(* Logix 5000 project; controller MV vendor 1 type 14 code 217 rev 31.11; software revision 31.00; part 46 of 53 *)
(* tags used below, declared in another part *)
   Always_Off : BOOL;
   CWD : CHECKWORD_FLAGS;
   Enable_TimeString : BOOL;
   MC_N100 : INT[255];   // C1_PLC Channel 1 PLC data
   MC_N120 : INT[255];   // C2 PLC Channel 2 PLC data
   MV_BM01_AV01 : PlantItem;   // BM01_AV01
   MV_BM01_AV01_CIP : BOOL;
   MV_BM01_AV01_mv22 : BOOL;
   MV_BM01_ZS04 : PlantItem;   // BM01ZS04
   MV_BM01_ZS05 : PlantItem;   // BM01ZS05
   MV_DAL01_AV01_mv22 : BOOL;
   MV_Data_To_TF : DINT[30];
   MV_Enable_MV22_NewPressureControl : BOOL;
   MV_FP01_ZS01 : PlantItem;   // FP01ZS01
   MV_FP01_ZS02 : PlantItem;   // FP01ZS02
   MV_GasAvailable : BOOL;
   MV_MV22_AV01 : PlantItem;   // MV22_AV01
   MV_MV22_CIP : BOOL;
   MV_MV22_CO2 : BOOL;
   MV_MV22_CO2_ON_PreStorage : BOOL;
   MV_MV22_CO2_ON_Storage : BOOL;
   MV_MV22_ControlOpenVent : BOOL;
   MV_MV22_Filling_Pulse : BOOL;
   MV_MV22_Filling_PulseLevel : DINT;
   MV_MV22_LTX07_TrueLevel : REAL;
   MV_MV22_ProxiesOK : BOOL;
   MV_MV22_PTX01_AI : PlantItem;   // MV22_PTX01
   MV_MV22_TP_CaskDepressure : BOOL;
   MV_MV22_TP_CaskEmptying : BOOL;
   MV_MV22_TP_CaskFilling : BOOL;
   MV_MV22_TP_CaskPreEmptyPressure : BOOL;
   MV_MV22_TP_CaskPrePressure : BOOL;
   MV_MV22_TP_CaskPressureDelay : BOOL;
   MV_MV22_TP_CaskReadyToFill : BOOL;
   MV_MV22_TP_CaskStorage : BOOL;
   MV_MV22_TP_CO2_Debounce_Timer : TIMER;
   MV_MV22_TP_CO2_Debounce_Timer_1 : TIMER;
   MV_MV22_TP_CO2_HSL_Pressure : REAL;
   MV_MV22_TP_CO2_HSL_Storage : REAL;
   MV_MV22_TP_CO2_HSL_Timer : TIMER;
   MV_MV22_TP_CO2_LSL_pressure_1 : REAL;
   MV_MV22_TP_CO2_LSL_storage : REAL;
   MV_MV22_TP_CO2_LSL_Timer : TIMER;
   MV_MV22_TP_Command : DINT;
   MV_MV22_TP_DAL_Chase_Cask : BOOL;
   MV_MV22_TP_DAL_Chase_KB : BOOL;
   MV_MV22_TP_DAL_Chase_Time : TIMER;
   MV_MV22_TP_Dirty : BOOL;
   MV_MV22_TP_Emptying_Level_Setpoint : REAL;
   MV_MV22_TP_Error_String : STRING;
   MV_MV22_TP_Faulted : BOOL;
   MV_MV22_TP_Fill_Pulse_OFF_Timer : TIMER;
   MV_MV22_TP_Fill_Pulse_ON_Timer : TIMER;
   MV_MV22_TP_Held : BOOL;
   MV_MV22_TP_Idle : BOOL;
   MV_MV22_TP_Initial_DAL_Chase_Cask : BOOL;
   MV_MV22_TP_Initial_DAL_Chase_KB : BOOL;
   MV_MV22_TP_KBEmptying : BOOL;
   MV_MV22_TP_KBFilling : BOOL;
   MV_MV22_TP_KBFillingBuildPressure : BOOL;
   MV_MV22_TP_KBPreEmptyPressure : BOOL;
   MV_MV22_TP_KBPrePressurise : BOOL;
   MV_MV22_TP_KBStorage : BOOL;
   MV_MV22_TP_LowerLimit : REAL;
   MV_MV22_TP_NotIdle : BOOL;
   MV_MV22_TP_ONS_1 : BOOL;
   MV_MV22_TP_Prompt : DINT;
   MV_MV22_TP_Proxy_Delay_Made : TIMER;
   MV_MV22_TP_Proxy_Delay_NOT_MADE : TIMER;
   MV_MV22_TP_Pulse : BOOL;
   MV_MV22_TP_ReadyToFillKB : BOOL;
   MV_MV22_TP_ReadyToFillKB_M : BOOL;
   MV_MV22_TP_Running : BOOL;
   MV_MV22_TP_Setpoint : REAL;
   MV_MV22_TP_Status : DINT;   // 0 = Idle, 1 = Running, 2 = Held, 3 = Faulted
   MV_MV22_TP_Step : DINT;
   MV_MV22_TP_Steptime : DINT;
   MV_MV22_TP_Steptime_String : STRING;
   MV_MV22_TP_SteptimeRunning : DINT;
   MV_MV22_TP_TimeLeft : DINT;
   MV_MV22_TP_TimeLeft_msec : DINT;
   MV_MV22_TP_TimeLeftStr : STRING;
   MV_MV22_TP_UpperLimit : REAL;
   MV_MV22_TP_Vent : BOOL;
   MV_MV22_TPLastStep : DINT;
   MV_N138 : INT[50];   // MV 22, CURRENT FV DATA
   MV_TP_CaskEmptyingPressure : REAL;
   MV_TP_CaskFillingPressure : REAL;
   MV_TP_CaskPrefillPressure : REAL;
   MV_TP_CaskStoragePressure : REAL;
   MV_TP_CaskStoragePressureDelay : DINT;
   MV_TP_CaskStoragePressureDelay_Secs : DINT;
   MV_TP_CaskStoragePressureLevel : REAL;
   MV_TP_Deadband : REAL;
   MV_TP_Emptying_Volume_Setpoint : REAL;
   MV_TP_HighLevelDeadband : REAL;
   MV_TP_KBFillingPressure : REAL;
   MV_TP_KBStoragePressure : REAL;
   MV_TP_LowLevelDeadbandThreshold : REAL;
   MV_TP_VentPressure : REAL;
   One_Second_1_scan : BOOL;
(* MV_Common, continued *)

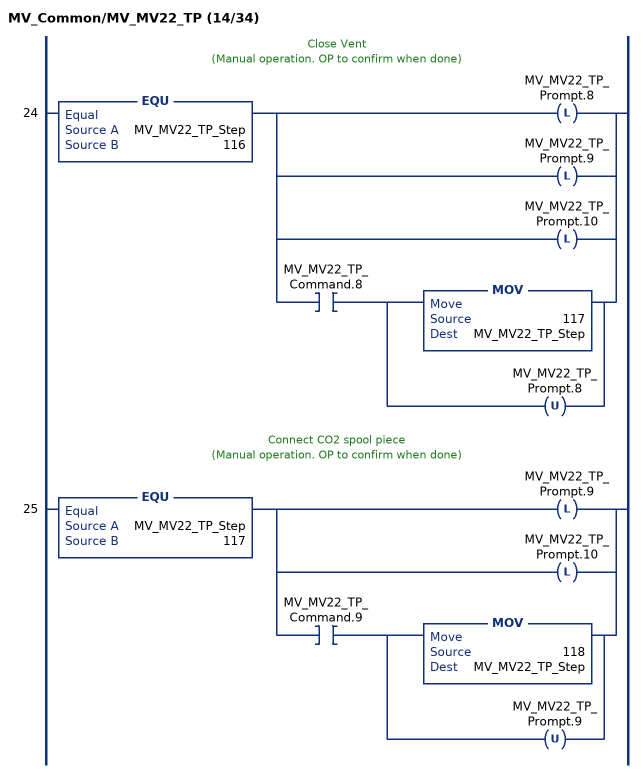
   // Close Vent
   // (Manual operation. OP to confirm when done)
   24: EQU(MV_MV22_TP_Step,116)[OTL(MV_MV22_TP_Prompt.8) ,OTL(MV_MV22_TP_Prompt.9) ,OTL(MV_MV22_TP_Prompt.10) ,XIC(MV_MV22_TP_Command.8) [MOV(117,MV_MV22_TP_Step) ,OTU(MV_MV22_TP_Prompt.8) ] ];
   // Connect CO2 spool piece
   // (Manual operation. OP to confirm when done)
   25: EQU(MV_MV22_TP_Step,117)[OTL(MV_MV22_TP_Prompt.9) ,OTL(MV_MV22_TP_Prompt.10) ,XIC(MV_MV22_TP_Command.9) [MOV(118,MV_MV22_TP_Step) ,OTU(MV_MV22_TP_Prompt.9) ] ];
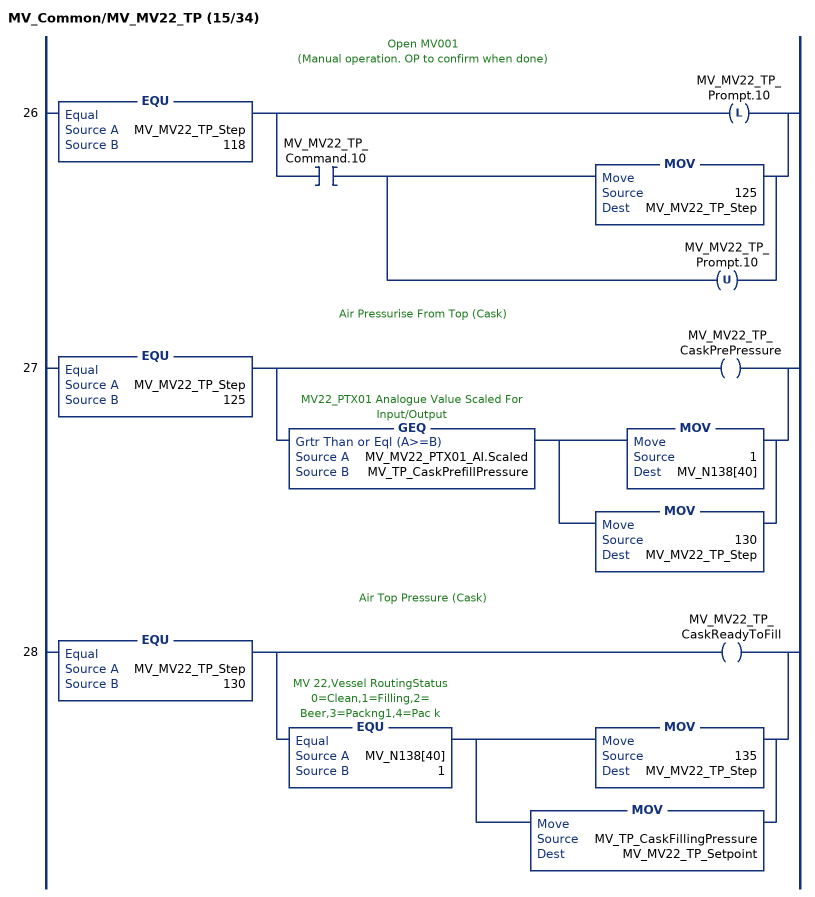
   // Open MV001
   // (Manual operation. OP to confirm when done)
   26: EQU(MV_MV22_TP_Step,118)[OTL(MV_MV22_TP_Prompt.10) ,XIC(MV_MV22_TP_Command.10) [MOV(125,MV_MV22_TP_Step) ,OTU(MV_MV22_TP_Prompt.10) ] ];
   // Air Pressurise From Top (Cask)
   27: EQU(MV_MV22_TP_Step,125)[OTE(MV_MV22_TP_CaskPrePressure) ,GEQ(MV_MV22_PTX01_AI.Scaled,MV_TP_CaskPrefillPressure) [MOV(1,MV_N138[40]) ,MOV(130,MV_MV22_TP_Step) ] ];
   // Air Top Pressure (Cask)
   28: EQU(MV_MV22_TP_Step,130)[OTE(MV_MV22_TP_CaskReadyToFill) ,EQU(MV_N138[40],1) [MOV(135,MV_MV22_TP_Step) ,MOV(MV_TP_CaskFillingPressure,MV_MV22_TP_Setpoint) ] ];
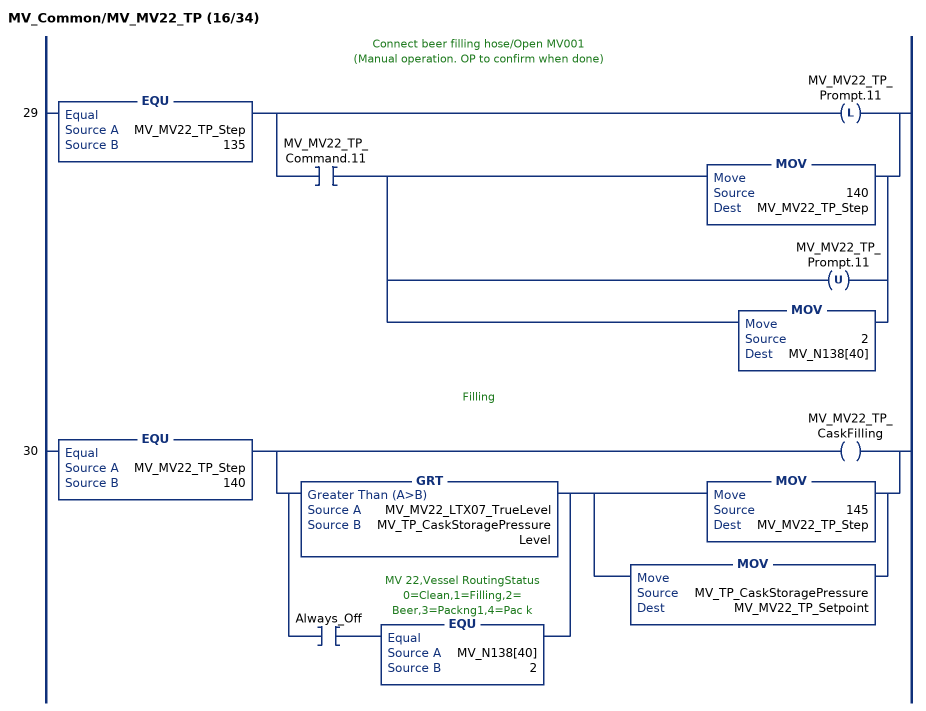
   // Connect beer filling hose/Open MV001
   // (Manual operation. OP to confirm when done)
   29: EQU(MV_MV22_TP_Step,135)[OTL(MV_MV22_TP_Prompt.11) ,XIC(MV_MV22_TP_Command.11) [MOV(140,MV_MV22_TP_Step) ,OTU(MV_MV22_TP_Prompt.11) ,MOV(2,MV_N138[40]) ] ];
   // Filling
   30: EQU(MV_MV22_TP_Step,140)[OTE(MV_MV22_TP_CaskFilling) ,[GRT(MV_MV22_LTX07_TrueLevel,MV_TP_CaskStoragePressureLevel) ,XIC(Always_Off) EQU(MV_N138[40],2) ] [MOV(145,MV_MV22_TP_Step) ,MOV(MV_TP_CaskStoragePressure,MV_MV22_TP_Setpoint) ] ];
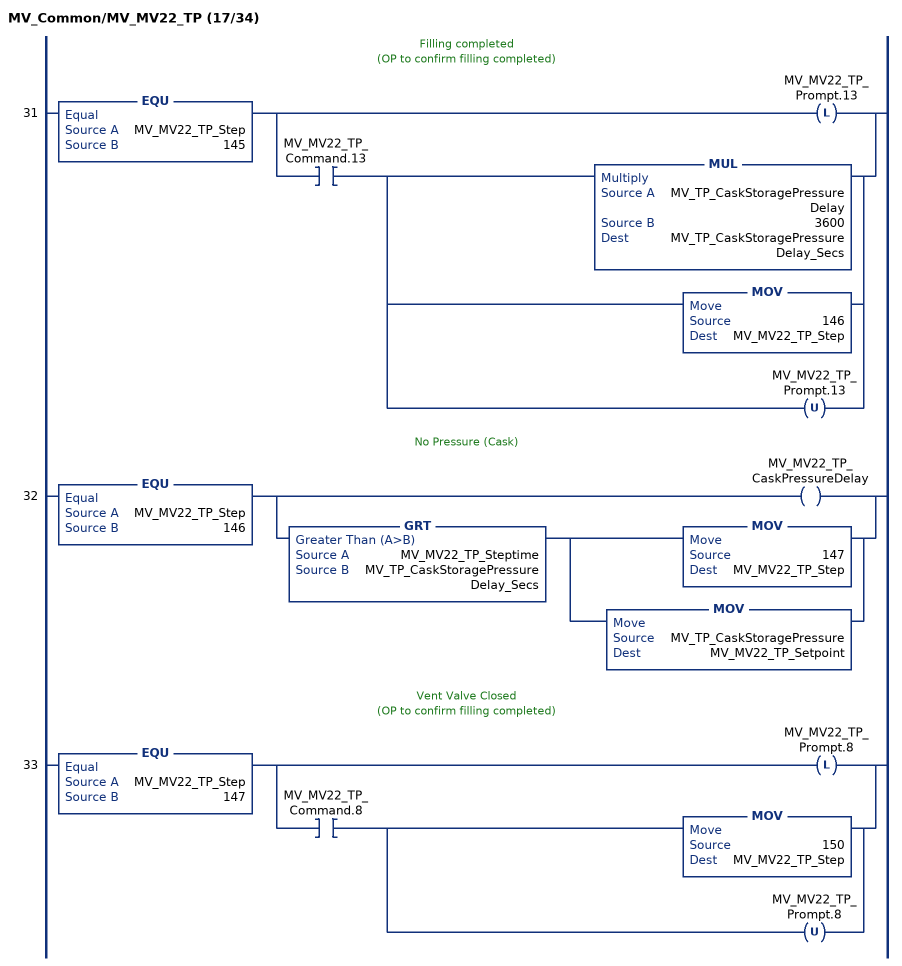
   // Filling completed
   // (OP to confirm filling completed)
   31: EQU(MV_MV22_TP_Step,145)[OTL(MV_MV22_TP_Prompt.13) ,XIC(MV_MV22_TP_Command.13) [MUL(MV_TP_CaskStoragePressureDelay,3600,MV_TP_CaskStoragePressureDelay_Secs) ,MOV(146,MV_MV22_TP_Step) ,OTU(MV_MV22_TP_Prompt.13) ] ];
   // No Pressure (Cask)
   32: EQU(MV_MV22_TP_Step,146)[OTE(MV_MV22_TP_CaskPressureDelay) ,GRT(MV_MV22_TP_Steptime,MV_TP_CaskStoragePressureDelay_Secs) [MOV(147,MV_MV22_TP_Step) ,MOV(MV_TP_CaskStoragePressure,MV_MV22_TP_Setpoint) ] ];
   // Vent Valve Closed
   // (OP to confirm filling completed)
   33: EQU(MV_MV22_TP_Step,147)[OTL(MV_MV22_TP_Prompt.8) ,XIC(MV_MV22_TP_Command.8) [MOV(150,MV_MV22_TP_Step) ,OTU(MV_MV22_TP_Prompt.8) ] ];
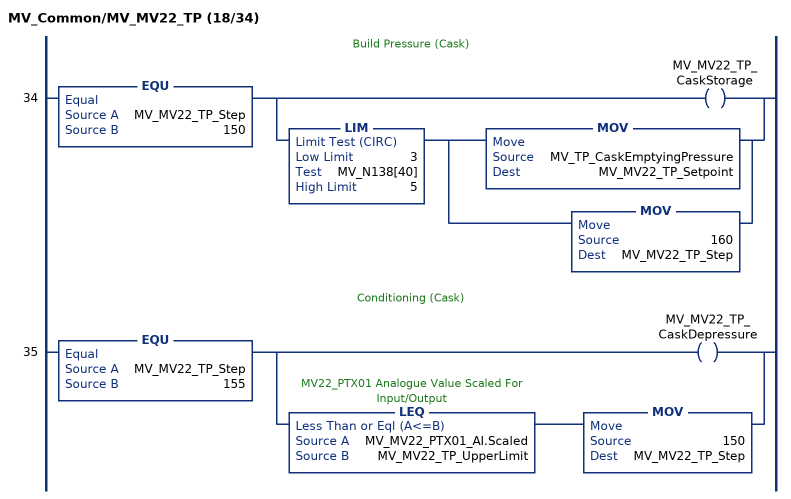
   // Build Pressure (Cask)
   34: EQU(MV_MV22_TP_Step,150)[OTE(MV_MV22_TP_CaskStorage) ,LIM(3,MV_N138[40],5) [MOV(MV_TP_CaskEmptyingPressure,MV_MV22_TP_Setpoint) ,MOV(160,MV_MV22_TP_Step) ] ];
   // Conditioning (Cask)
   35: EQU(MV_MV22_TP_Step,155)[OTE(MV_MV22_TP_CaskDepressure) ,LEQ(MV_MV22_PTX01_AI.Scaled,MV_MV22_TP_UpperLimit) MOV(150,MV_MV22_TP_Step) ];
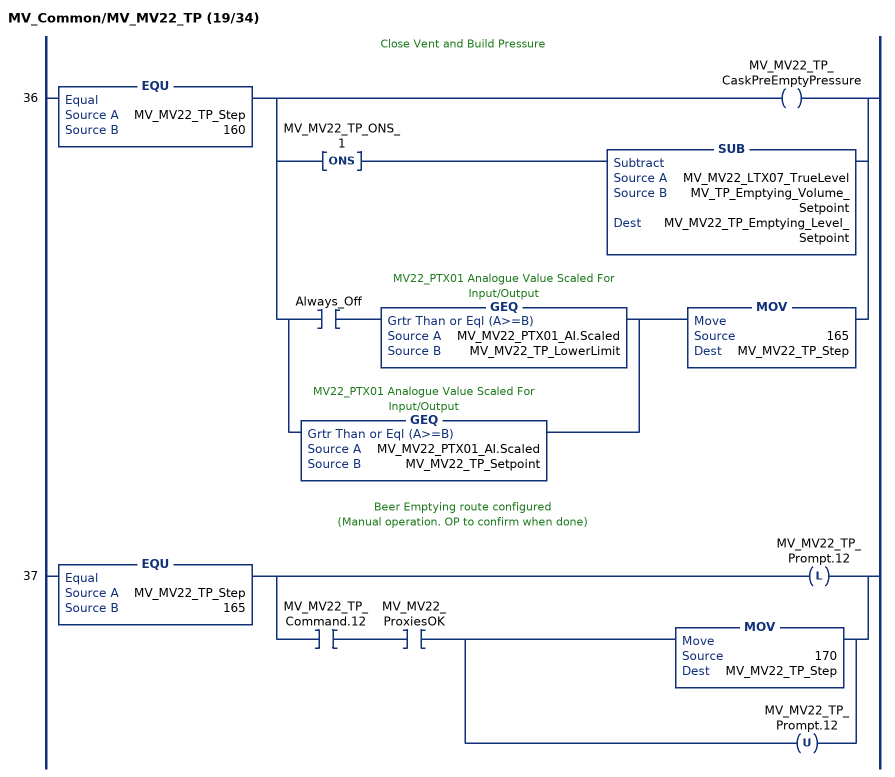
   // Close Vent and Build Pressure
   36: EQU(MV_MV22_TP_Step,160)[OTE(MV_MV22_TP_CaskPreEmptyPressure) ,ONS(MV_MV22_TP_ONS_1) SUB(MV_MV22_LTX07_TrueLevel,MV_TP_Emptying_Volume_Setpoint,MV_MV22_TP_Emptying_Level_Setpoint) ,[XIC(Always_Off) GEQ(MV_MV22_PTX01_AI.Scaled,MV_MV22_TP_LowerLimit) ,GEQ(MV_MV22_PTX01_AI.Scaled,MV_MV22_TP_Setpoint) ] MOV(165,MV_MV22_TP_Step) ];
   // Beer Emptying route configured
   // (Manual operation. OP to confirm when done)
   37: EQU(MV_MV22_TP_Step,165)[OTL(MV_MV22_TP_Prompt.12) ,XIC(MV_MV22_TP_Command.12) XIC(MV_MV22_ProxiesOK) [MOV(170,MV_MV22_TP_Step) ,OTU(MV_MV22_TP_Prompt.12) ] ];
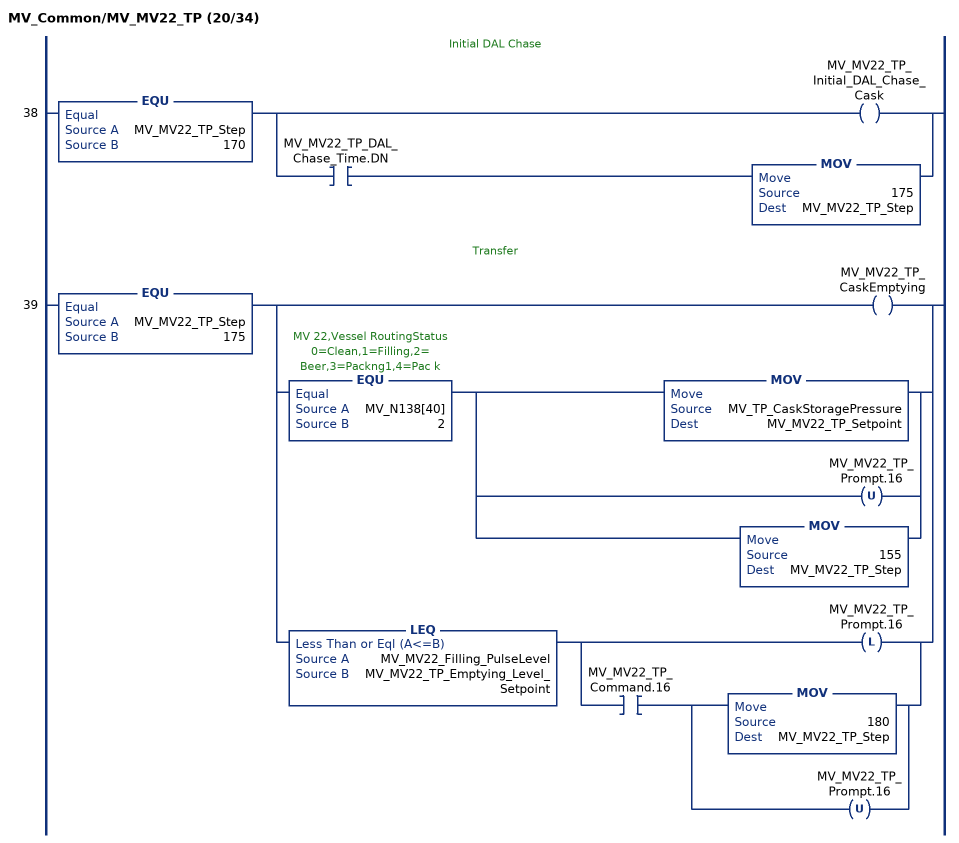
   // Initial DAL Chase
   38: EQU(MV_MV22_TP_Step,170)[OTE(MV_MV22_TP_Initial_DAL_Chase_Cask) ,XIC(MV_MV22_TP_DAL_Chase_Time.DN) MOV(175,MV_MV22_TP_Step) ];
   // Transfer
   39: EQU(MV_MV22_TP_Step,175)[OTE(MV_MV22_TP_CaskEmptying) ,EQU(MV_N138[40],2) [MOV(MV_TP_CaskStoragePressure,MV_MV22_TP_Setpoint) ,OTU(MV_MV22_TP_Prompt.16) ,MOV(155,MV_MV22_TP_Step) ] ,LEQ(MV_MV22_Filling_PulseLevel,MV_MV22_TP_Emptying_Level_Setpoint) [OTL(MV_MV22_TP_Prompt.16) ,XIC(MV_MV22_TP_Command.16) [MOV(180,MV_MV22_TP_Step) ,OTU(MV_MV22_TP_Prompt.16) ] ] ];
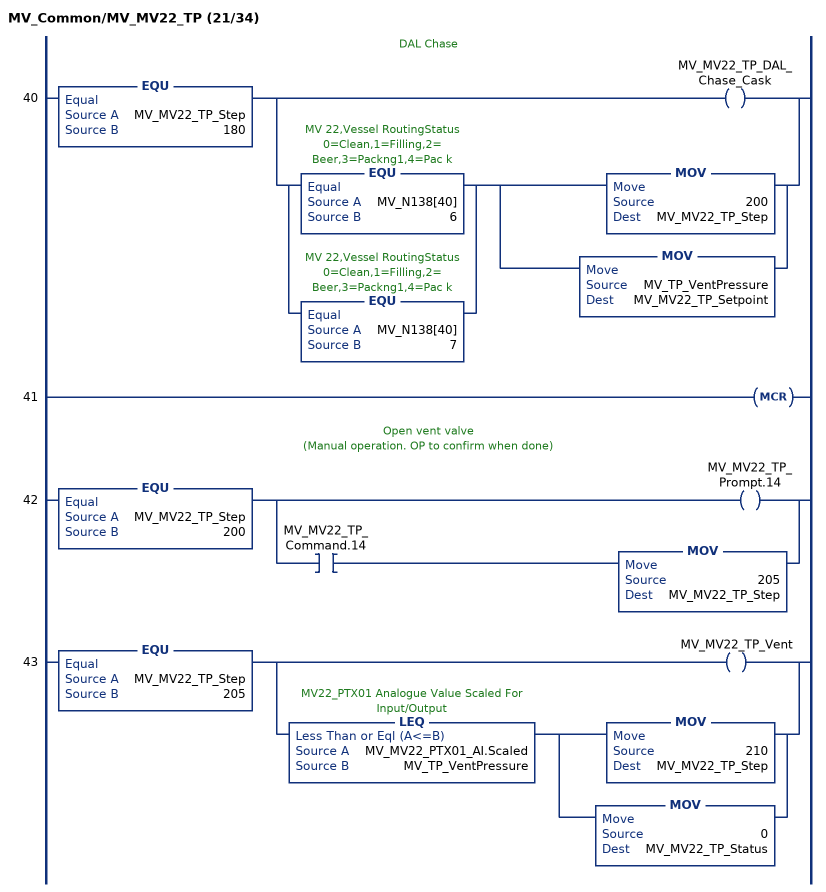
   // DAL Chase
   40: EQU(MV_MV22_TP_Step,180)[OTE(MV_MV22_TP_DAL_Chase_Cask) ,[EQU(MV_N138[40],6) ,EQU(MV_N138[40],7) ] [MOV(200,MV_MV22_TP_Step) ,MOV(MV_TP_VentPressure,MV_MV22_TP_Setpoint) ] ];
   41: MCR();
   // Open vent valve
   // (Manual operation. OP to confirm when done)
   42: EQU(MV_MV22_TP_Step,200)[OTE(MV_MV22_TP_Prompt.14) ,XIC(MV_MV22_TP_Command.14) MOV(205,MV_MV22_TP_Step) ];
   43: EQU(MV_MV22_TP_Step,205)[OTE(MV_MV22_TP_Vent) ,LEQ(MV_MV22_PTX01_AI.Scaled,MV_TP_VentPressure) [MOV(210,MV_MV22_TP_Step) ,MOV(0,MV_MV22_TP_Status) ] ];
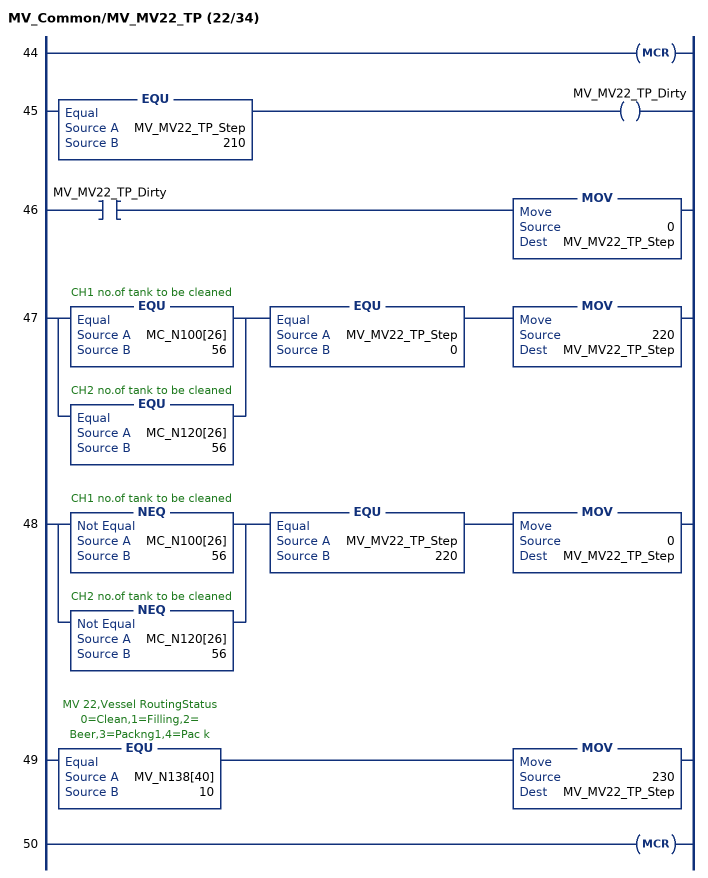
   44: MCR();
   45: EQU(MV_MV22_TP_Step,210)OTE(MV_MV22_TP_Dirty);
   46: XIC(MV_MV22_TP_Dirty)MOV(0,MV_MV22_TP_Step);
   47: [EQU(MC_N100[26],56) ,EQU(MC_N120[26],56) ]EQU(MV_MV22_TP_Step,0)MOV(220,MV_MV22_TP_Step);
   48: [NEQ(MC_N100[26],56) ,NEQ(MC_N120[26],56) ]EQU(MV_MV22_TP_Step,220)MOV(0,MV_MV22_TP_Step);
   49: EQU(MV_N138[40],10)MOV(230,MV_MV22_TP_Step);
   50: MCR();
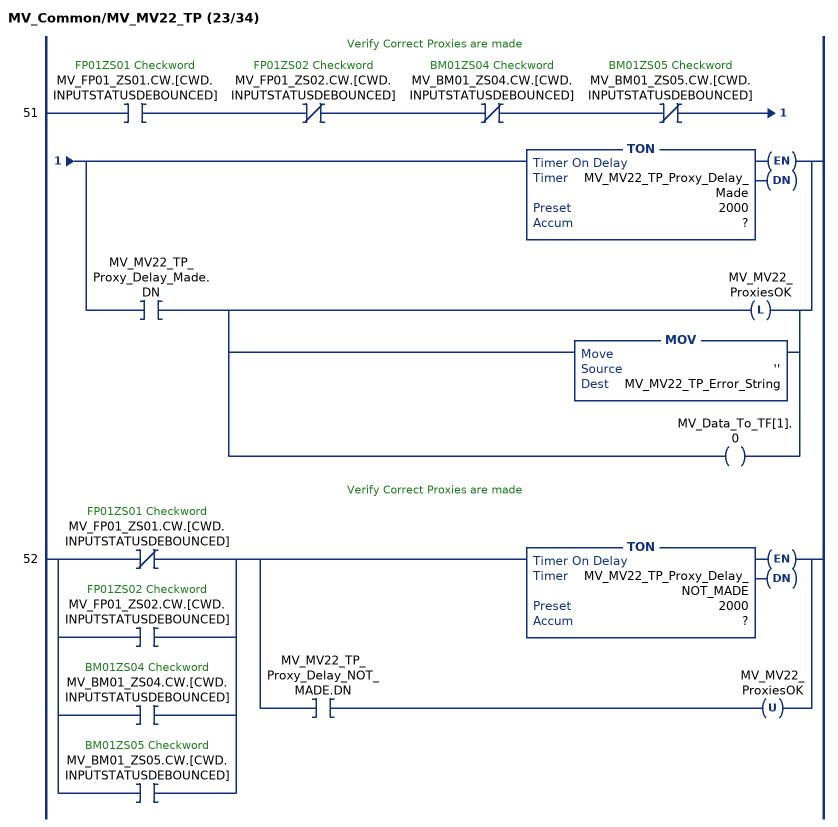
   // Verify Correct Proxies are made
   51: XIC(MV_FP01_ZS01.CW.[CWD.INPUTSTATUSDEBOUNCED])XIO(MV_FP01_ZS02.CW.[CWD.INPUTSTATUSDEBOUNCED])XIO(MV_BM01_ZS04.CW.[CWD.INPUTSTATUSDEBOUNCED])XIO(MV_BM01_ZS05.CW.[CWD.INPUTSTATUSDEBOUNCED])[TON(MV_MV22_TP_Proxy_Delay_Made,?,?) ,XIC(MV_MV22_TP_Proxy_Delay_Made.DN) [OTL(MV_MV22_ProxiesOK) ,MOV('',MV_MV22_TP_Error_String) ,OTE(MV_Data_To_TF[1].0) ] ];
   // Verify Correct Proxies are made
   52: [XIO(MV_FP01_ZS01.CW.[CWD.INPUTSTATUSDEBOUNCED]) ,XIC(MV_FP01_ZS02.CW.[CWD.INPUTSTATUSDEBOUNCED]) ,XIC(MV_BM01_ZS04.CW.[CWD.INPUTSTATUSDEBOUNCED]) ,XIC(MV_BM01_ZS05.CW.[CWD.INPUTSTATUSDEBOUNCED]) ][TON(MV_MV22_TP_Proxy_Delay_NOT_MADE,?,?) ,XIC(MV_MV22_TP_Proxy_Delay_NOT_MADE.DN) OTU(MV_MV22_ProxiesOK) ];
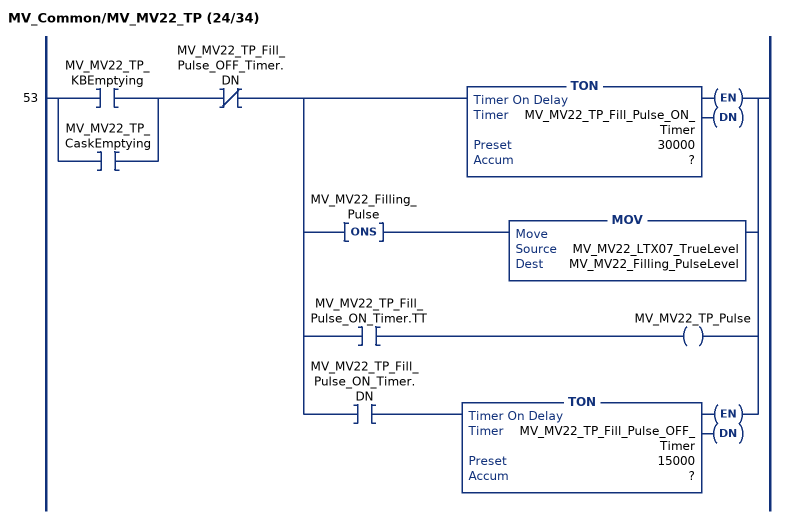
   53: [XIC(MV_MV22_TP_KBEmptying) ,XIC(MV_MV22_TP_CaskEmptying) ]XIO(MV_MV22_TP_Fill_Pulse_OFF_Timer.DN)[TON(MV_MV22_TP_Fill_Pulse_ON_Timer,?,?) ,ONS(MV_MV22_Filling_Pulse) MOV(MV_MV22_LTX07_TrueLevel,MV_MV22_Filling_PulseLevel) ,XIC(MV_MV22_TP_Fill_Pulse_ON_Timer.TT) OTE(MV_MV22_TP_Pulse) ,XIC(MV_MV22_TP_Fill_Pulse_ON_Timer.DN) TON(MV_MV22_TP_Fill_Pulse_OFF_Timer,?,?) ];
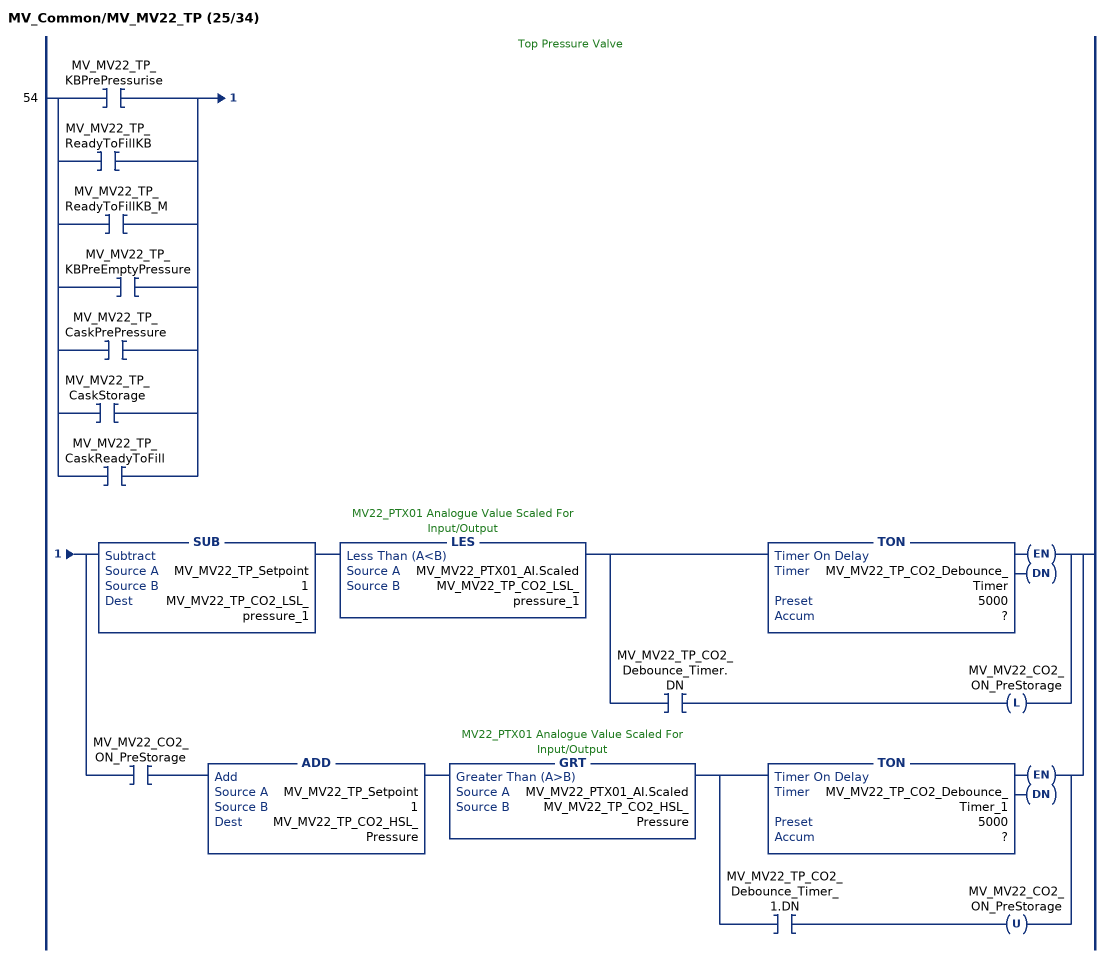
   // Top Pressure Valve
   54: [XIC(MV_MV22_TP_KBPrePressurise) ,XIC(MV_MV22_TP_ReadyToFillKB) ,XIC(MV_MV22_TP_ReadyToFillKB_M) ,XIC(MV_MV22_TP_KBPreEmptyPressure) ,XIC(MV_MV22_TP_CaskPrePressure) ,XIC(MV_MV22_TP_CaskStorage) ,XIC(MV_MV22_TP_CaskReadyToFill) ][SUB(MV_MV22_TP_Setpoint,1,MV_MV22_TP_CO2_LSL_pressure_1) LES(MV_MV22_PTX01_AI.Scaled,MV_MV22_TP_CO2_LSL_pressure_1) [TON(MV_MV22_TP_CO2_Debounce_Timer,?,?) ,XIC(MV_MV22_TP_CO2_Debounce_Timer.DN) OTL(MV_MV22_CO2_ON_PreStorage) ] ,XIC(MV_MV22_CO2_ON_PreStorage) ADD(MV_MV22_TP_Setpoint,1,MV_MV22_TP_CO2_HSL_Pressure) GRT(MV_MV22_PTX01_AI.Scaled,MV_MV22_TP_CO2_HSL_Pressure) [TON(MV_MV22_TP_CO2_Debounce_Timer_1,?,?) ,XIC(MV_MV22_TP_CO2_Debounce_Timer_1.DN) OTU(MV_MV22_CO2_ON_PreStorage) ] ];
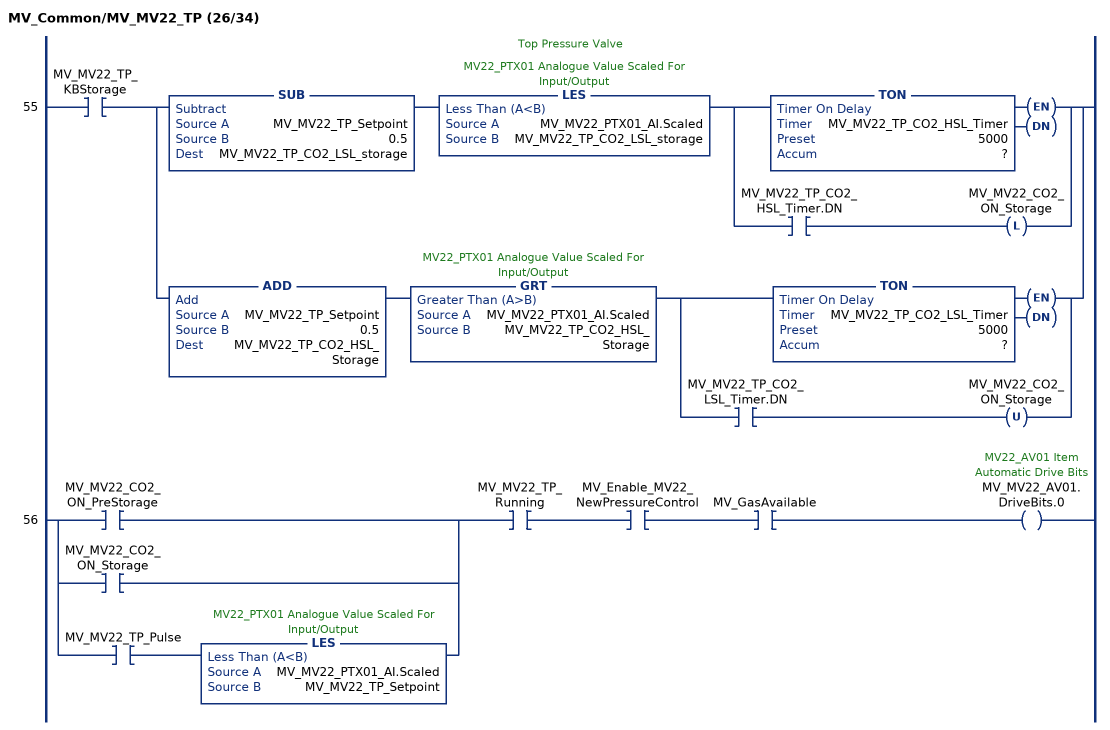
   // Top Pressure Valve
   55: XIC(MV_MV22_TP_KBStorage)[SUB(MV_MV22_TP_Setpoint,0.5,MV_MV22_TP_CO2_LSL_storage) LES(MV_MV22_PTX01_AI.Scaled,MV_MV22_TP_CO2_LSL_storage) [TON(MV_MV22_TP_CO2_HSL_Timer,?,?) ,XIC(MV_MV22_TP_CO2_HSL_Timer.DN) OTL(MV_MV22_CO2_ON_Storage) ] ,ADD(MV_MV22_TP_Setpoint,0.5,MV_MV22_TP_CO2_HSL_Storage) GRT(MV_MV22_PTX01_AI.Scaled,MV_MV22_TP_CO2_HSL_Storage) [TON(MV_MV22_TP_CO2_LSL_Timer,?,?) ,XIC(MV_MV22_TP_CO2_LSL_Timer.DN) OTU(MV_MV22_CO2_ON_Storage) ] ];
   56: [XIC(MV_MV22_CO2_ON_PreStorage) ,XIC(MV_MV22_CO2_ON_Storage) ,XIC(MV_MV22_TP_Pulse) LES(MV_MV22_PTX01_AI.Scaled,MV_MV22_TP_Setpoint) ]XIC(MV_MV22_TP_Running)XIC(MV_Enable_MV22_NewPressureControl)XIC(MV_GasAvailable)OTE(MV_MV22_AV01.DriveBits.0);
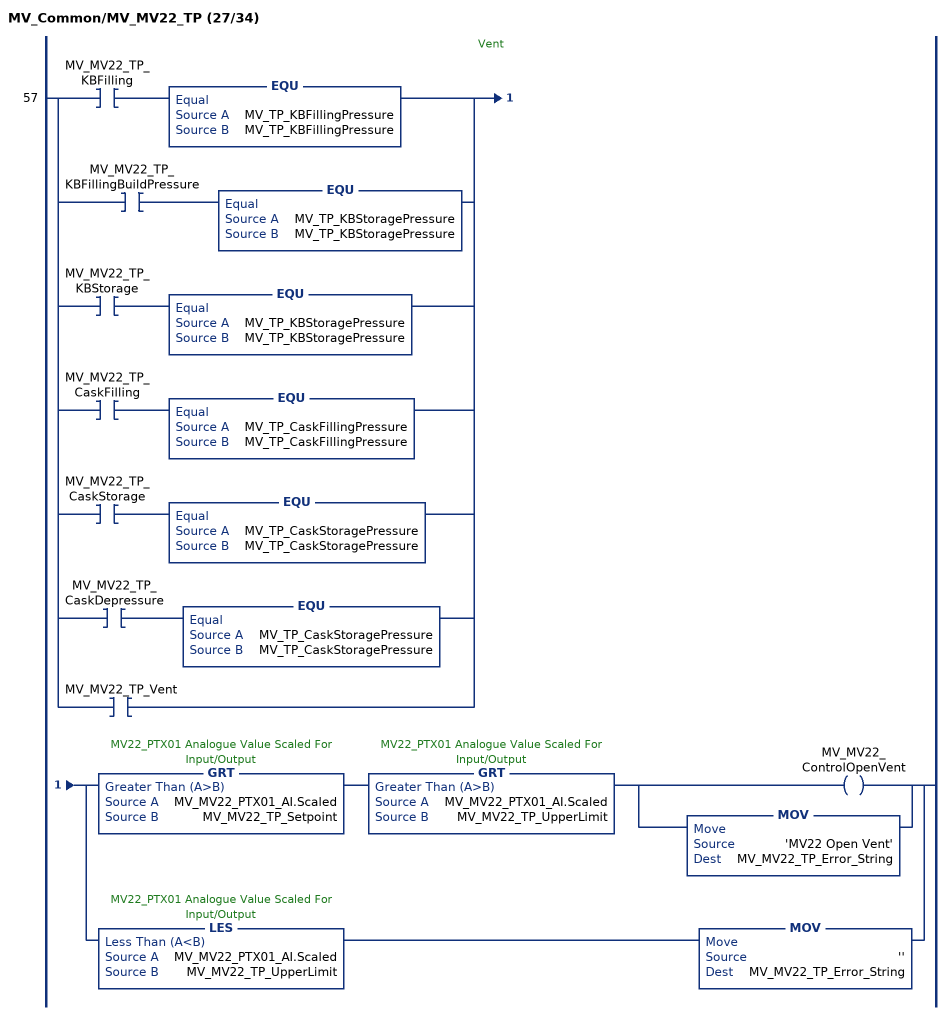
   // Vent
   57: [XIC(MV_MV22_TP_KBFilling) EQU(MV_TP_KBFillingPressure,MV_TP_KBFillingPressure) ,XIC(MV_MV22_TP_KBFillingBuildPressure) EQU(MV_TP_KBStoragePressure,MV_TP_KBStoragePressure) ,XIC(MV_MV22_TP_KBStorage) EQU(MV_TP_KBStoragePressure,MV_TP_KBStoragePressure) ,XIC(MV_MV22_TP_CaskFilling) EQU(MV_TP_CaskFillingPressure,MV_TP_CaskFillingPressure) ,XIC(MV_MV22_TP_CaskStorage) EQU(MV_TP_CaskStoragePressure,MV_TP_CaskStoragePressure) ,XIC(MV_MV22_TP_CaskDepressure) EQU(MV_TP_CaskStoragePressure,MV_TP_CaskStoragePressure) ,XIC(MV_MV22_TP_Vent) ][GRT(MV_MV22_PTX01_AI.Scaled,MV_MV22_TP_Setpoint) GRT(MV_MV22_PTX01_AI.Scaled,MV_MV22_TP_UpperLimit) [OTE(MV_MV22_ControlOpenVent) ,MOV('MV22 Open Vent',MV_MV22_TP_Error_String) ] ,LES(MV_MV22_PTX01_AI.Scaled,MV_MV22_TP_UpperLimit) MOV('',MV_MV22_TP_Error_String) ];
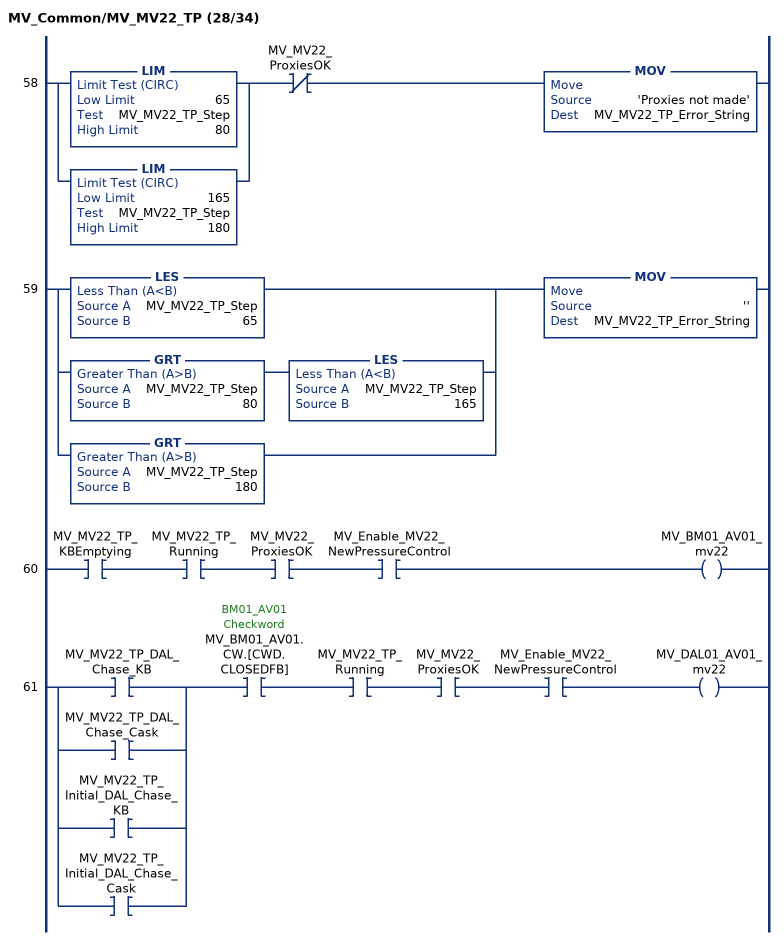
   58: [LIM(65,MV_MV22_TP_Step,80) ,LIM(165,MV_MV22_TP_Step,180) ]XIO(MV_MV22_ProxiesOK)MOV('Proxies not made',MV_MV22_TP_Error_String);
   59: [LES(MV_MV22_TP_Step,65) ,GRT(MV_MV22_TP_Step,80) LES(MV_MV22_TP_Step,165) ,GRT(MV_MV22_TP_Step,180) ]MOV('',MV_MV22_TP_Error_String);
   60: XIC(MV_MV22_TP_KBEmptying)XIC(MV_MV22_TP_Running)XIC(MV_MV22_ProxiesOK)XIC(MV_Enable_MV22_NewPressureControl)OTE(MV_BM01_AV01_mv22);
   61: [XIC(MV_MV22_TP_DAL_Chase_KB) ,XIC(MV_MV22_TP_DAL_Chase_Cask) ,XIC(MV_MV22_TP_Initial_DAL_Chase_KB) ,XIC(MV_MV22_TP_Initial_DAL_Chase_Cask) ]XIC(MV_BM01_AV01.CW.[CWD.CLOSEDFB])XIC(MV_MV22_TP_Running)XIC(MV_MV22_ProxiesOK)XIC(MV_Enable_MV22_NewPressureControl)OTE(MV_DAL01_AV01_mv22);
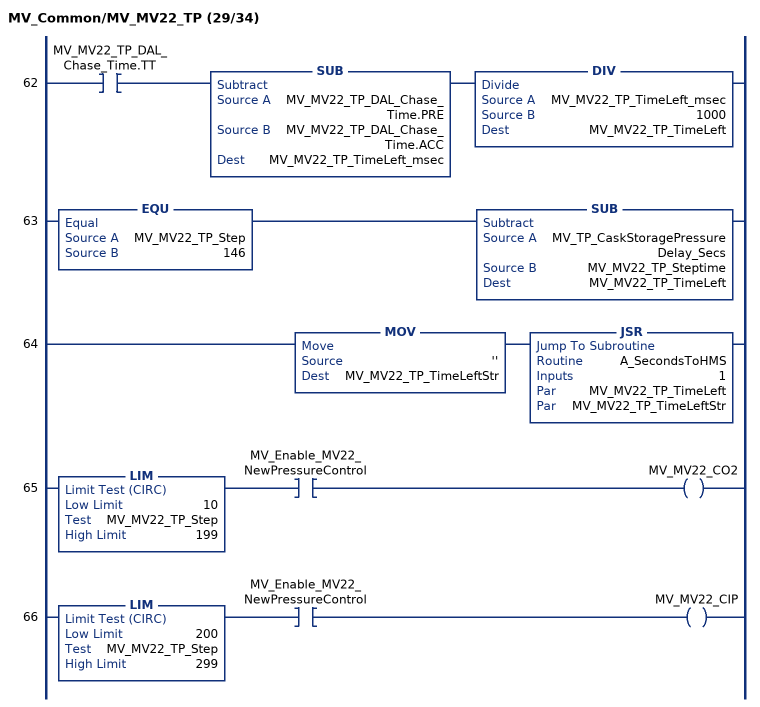
   62: XIC(MV_MV22_TP_DAL_Chase_Time.TT)SUB(MV_MV22_TP_DAL_Chase_Time.PRE,MV_MV22_TP_DAL_Chase_Time.ACC,MV_MV22_TP_TimeLeft_msec)DIV(MV_MV22_TP_TimeLeft_msec,1000,MV_MV22_TP_TimeLeft);
   63: EQU(MV_MV22_TP_Step,146)SUB(MV_TP_CaskStoragePressureDelay_Secs,MV_MV22_TP_Steptime,MV_MV22_TP_TimeLeft);
   64: MOV('',MV_MV22_TP_TimeLeftStr)JSR(A_SecondsToHMS,1,MV_MV22_TP_TimeLeft,MV_MV22_TP_TimeLeftStr);
   65: LIM(10,MV_MV22_TP_Step,199)XIC(MV_Enable_MV22_NewPressureControl)OTE(MV_MV22_CO2);
   66: LIM(200,MV_MV22_TP_Step,299)XIC(MV_Enable_MV22_NewPressureControl)OTE(MV_MV22_CIP);
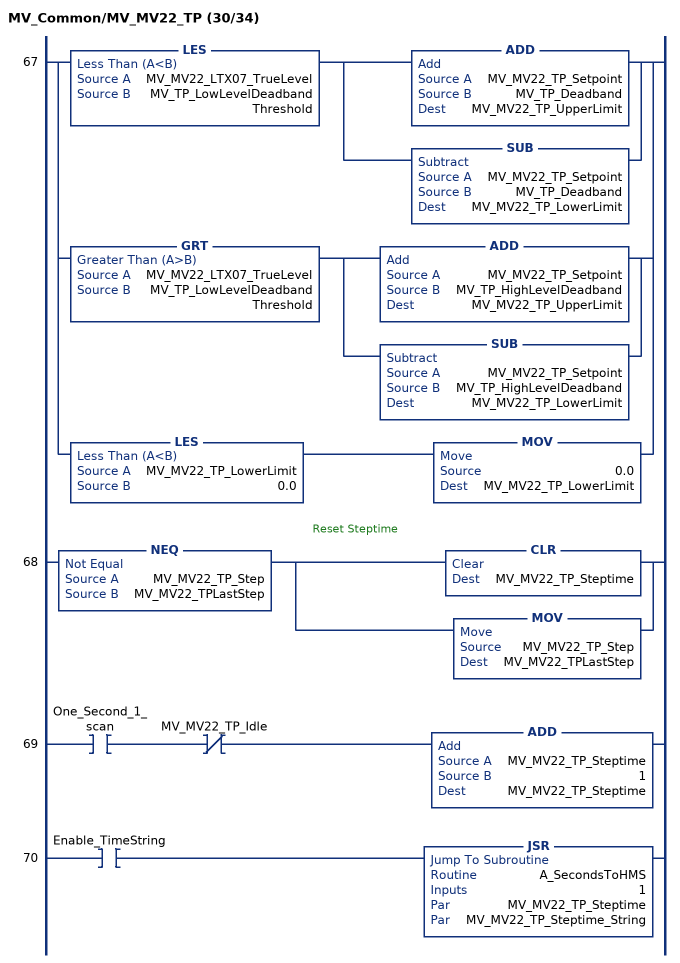
   67: [LES(MV_MV22_LTX07_TrueLevel,MV_TP_LowLevelDeadbandThreshold) [ADD(MV_MV22_TP_Setpoint,MV_TP_Deadband,MV_MV22_TP_UpperLimit) ,SUB(MV_MV22_TP_Setpoint,MV_TP_Deadband,MV_MV22_TP_LowerLimit) ] ,GRT(MV_MV22_LTX07_TrueLevel,MV_TP_LowLevelDeadbandThreshold) [ADD(MV_MV22_TP_Setpoint,MV_TP_HighLevelDeadband,MV_MV22_TP_UpperLimit) ,SUB(MV_MV22_TP_Setpoint,MV_TP_HighLevelDeadband,MV_MV22_TP_LowerLimit) ] ,LES(MV_MV22_TP_LowerLimit,0.0) MOV(0.0,MV_MV22_TP_LowerLimit) ];
   // Reset Steptime
   68: NEQ(MV_MV22_TP_Step,MV_MV22_TPLastStep)[CLR(MV_MV22_TP_Steptime) ,MOV(MV_MV22_TP_Step,MV_MV22_TPLastStep) ];
   69: XIC(One_Second_1_scan)XIO(MV_MV22_TP_Idle)ADD(MV_MV22_TP_Steptime,1,MV_MV22_TP_Steptime);
   70: XIC(Enable_TimeString)JSR(A_SecondsToHMS,1,MV_MV22_TP_Steptime,MV_MV22_TP_Steptime_String);
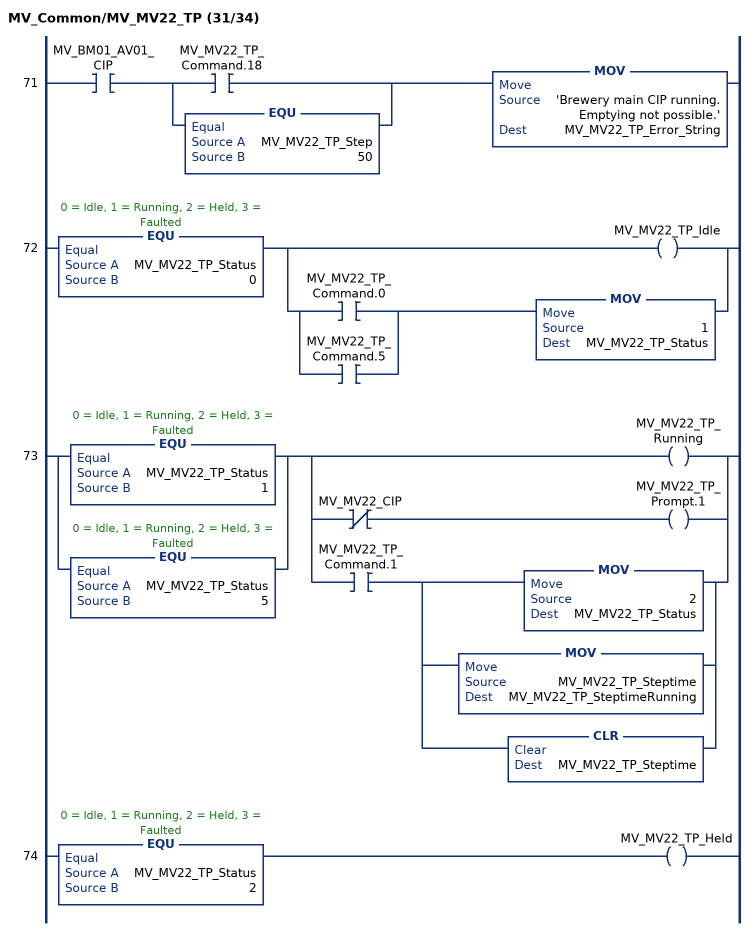
   71: XIC(MV_BM01_AV01_CIP)[XIC(MV_MV22_TP_Command.18) ,EQU(MV_MV22_TP_Step,50) ]MOV('Brewery main CIP running. Emptying not possible.',MV_MV22_TP_Error_String);
   72: EQU(MV_MV22_TP_Status,0)[OTE(MV_MV22_TP_Idle) ,[XIC(MV_MV22_TP_Command.0) ,XIC(MV_MV22_TP_Command.5) ] MOV(1,MV_MV22_TP_Status) ];
   73: [EQU(MV_MV22_TP_Status,1) ,EQU(MV_MV22_TP_Status,5) ][OTE(MV_MV22_TP_Running) ,XIO(MV_MV22_CIP) OTE(MV_MV22_TP_Prompt.1) ,XIC(MV_MV22_TP_Command.1) [MOV(2,MV_MV22_TP_Status) ,MOV(MV_MV22_TP_Steptime,MV_MV22_TP_SteptimeRunning) ,CLR(MV_MV22_TP_Steptime) ] ];
   74: EQU(MV_MV22_TP_Status,2)OTE(MV_MV22_TP_Held);
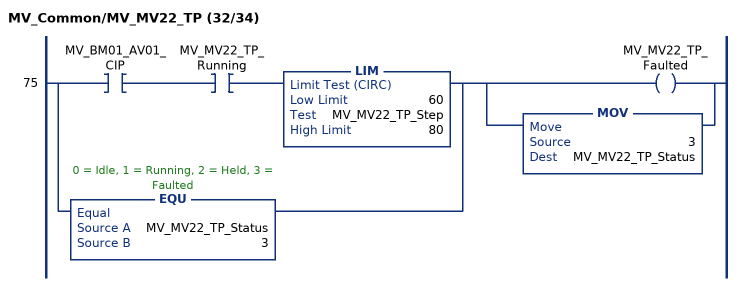
   75: [XIC(MV_BM01_AV01_CIP) XIC(MV_MV22_TP_Running) LIM(60,MV_MV22_TP_Step,80) ,EQU(MV_MV22_TP_Status,3) ][OTE(MV_MV22_TP_Faulted) ,MOV(3,MV_MV22_TP_Status) ];
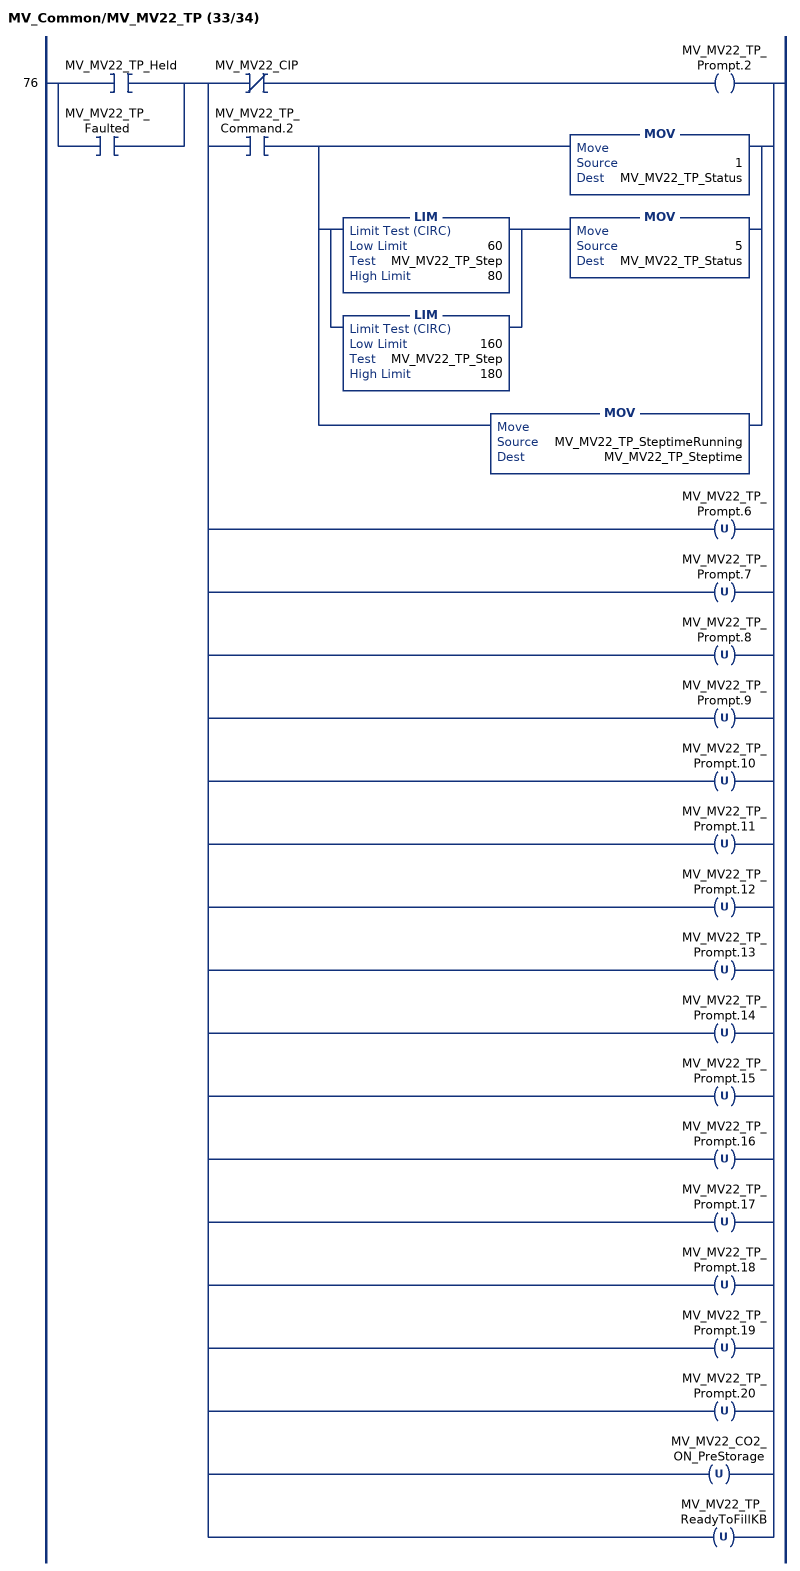
   76: [XIC(MV_MV22_TP_Held) ,XIC(MV_MV22_TP_Faulted) ][XIO(MV_MV22_CIP) OTE(MV_MV22_TP_Prompt.2) ,XIC(MV_MV22_TP_Command.2) [MOV(1,MV_MV22_TP_Status) ,[LIM(60,MV_MV22_TP_Step,80) ,LIM(160,MV_MV22_TP_Step,180) ] MOV(5,MV_MV22_TP_Status) ,MOV(MV_MV22_TP_SteptimeRunning,MV_MV22_TP_Steptime) ] ,OTU(MV_MV22_TP_Prompt.6) ,OTU(MV_MV22_TP_Prompt.7) ,OTU(MV_MV22_TP_Prompt.8) ,OTU(MV_MV22_TP_Prompt.9) ,OTU(MV_MV22_TP_Prompt.10) ,OTU(MV_MV22_TP_Prompt.11) ,OTU(MV_MV22_TP_Prompt.12) ,OTU(MV_MV22_TP_Prompt.13) ,OTU(MV_MV22_TP_Prompt.14) ,OTU(MV_MV22_TP_Prompt.15) ,OTU(MV_MV22_TP_Prompt.16) ,OTU(MV_MV22_TP_Prompt.17) ,OTU(MV_MV22_TP_Prompt.18) ,OTU(MV_MV22_TP_Prompt.19) ,OTU(MV_MV22_TP_Prompt.20) ,OTU(MV_MV22_CO2_ON_PreStorage) ,OTU(MV_MV22_TP_ReadyToFillKB) ];
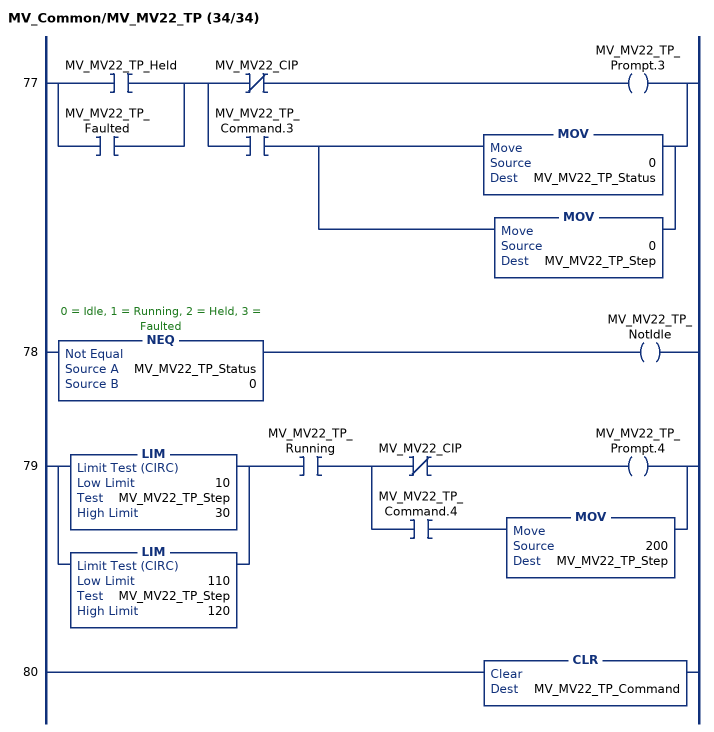
   77: [XIC(MV_MV22_TP_Held) ,XIC(MV_MV22_TP_Faulted) ][XIO(MV_MV22_CIP) OTE(MV_MV22_TP_Prompt.3) ,XIC(MV_MV22_TP_Command.3) [MOV(0,MV_MV22_TP_Status) ,MOV(0,MV_MV22_TP_Step) ] ];
   78: NEQ(MV_MV22_TP_Status,0)OTE(MV_MV22_TP_NotIdle);
   79: [LIM(10,MV_MV22_TP_Step,30) ,LIM(110,MV_MV22_TP_Step,120) ]XIC(MV_MV22_TP_Running)[XIO(MV_MV22_CIP) OTE(MV_MV22_TP_Prompt.4) ,XIC(MV_MV22_TP_Command.4) MOV(200,MV_MV22_TP_Step) ];
   80: CLR(MV_MV22_TP_Command);
END_ROUTINE
